(* Logix 5000 project; controller MV vendor 1 type 14 code 217 rev 31.11; software revision 31.00; part 30 of 53 *)
(* tags used below, declared in another part *)
   Alarm_Reset : BOOL;
   CWD : CHECKWORD_FLAGS;
   Default_Check_Time : DINT;
   Item_Faults_Are_Latched : BOOL;
   Item_Simulation_Flag : BOOL;
   MC_CH1_DR1 : PlantItem;   // CH1_DR1
   MC_CH1_DR1_ALARM : ALARM_DIGITAL;
   MC_CH1_DR1_C : ALIAS FOR RIO_Rack_2:4:I.Data.30;
   MC_CH1_DR1_DR : ALIAS FOR RIO_Rack_2:5:O.Data.14;
   MC_CH1_DR1_O : ALIAS FOR RIO_Rack_2:4:I.Data.26;
   MC_CH1_DR2 : PlantItem;   // CH1_DR2
   MC_CH1_DR2_ALARM : ALARM_DIGITAL;
   MC_CH1_DR2_C : ALIAS FOR RIO_Rack_2:4:I.Data.31;
   MC_CH1_DR2_DR : ALIAS FOR RIO_Rack_2:5:O.Data.15;
   MC_CH1_DR2_O : ALIAS FOR RIO_Rack_2:4:I.Data.27;
   MC_CH1_DRAIN : PlantItem;   // CH1_DRAIN
   MC_CH1_DRAIN_ALARM : ALARM_DIGITAL;
   MC_CH1_DRAIN_C : ALIAS FOR RIO_Rack_2:4:I.Data.28;
   MC_CH1_DRAIN_DR : ALIAS FOR RIO_Rack_2:5:O.Data.12;
   MC_CH1_DRAIN_O : ALIAS FOR RIO_Rack_2:4:I.Data.24;
   MC_CH1_DT1 : PlantItem;   // CH1_DT1
   MC_CH1_DT1_ALARM : ALARM_DIGITAL;
   MC_CH1_DT1_C : ALIAS FOR RIO_Rack_2:6:I.Data.4;
   MC_CH1_DT1_DR : ALIAS FOR RIO_Rack_2:5:O.Data.16;
   MC_CH1_DT1_O : ALIAS FOR RIO_Rack_2:6:I.Data.0;
   MC_CH1_DT2 : PlantItem;   // CH1_DT2
   MC_CH1_DT2_ALARM : ALARM_DIGITAL;
   MC_CH1_DT2_C : ALIAS FOR RIO_Rack_2:6:I.Data.5;
   MC_CH1_DT2_DR : ALIAS FOR RIO_Rack_2:5:O.Data.17;
   MC_CH1_DT2_O : ALIAS FOR RIO_Rack_2:6:I.Data.1;
   MC_CH1_LF1 : PlantItem;   // CH1_LF1
   MC_CH1_LF1_ALARM : ALARM_DIGITAL;
   MC_CH1_LF1_C : ALIAS FOR RIO_Rack_2:6:I.Data.7;
   MC_CH1_LF1_DR : ALIAS FOR RIO_Rack_2:5:O.Data.19;
   MC_CH1_LF1_O : ALIAS FOR RIO_Rack_2:6:I.Data.3;
   MC_CH1_PR1 : PlantItem;   // CH1_PR1
   MC_CH1_PR1_ALARM : ALARM_DIGITAL;
   MC_CH1_PR1_C : ALIAS FOR RIO_Rack_2:6:I.Data.6;
   MC_CH1_PR1_DR : ALIAS FOR RIO_Rack_2:5:O.Data.18;
   MC_CH1_PR1_O : ALIAS FOR RIO_Rack_2:6:I.Data.2;
   MC_CH1_R2R : PlantItem;   // CH1_R2R
   MC_CH1_R2R_ALARM : ALARM_DIGITAL;
   MC_CH1_R2R_C : ALIAS FOR RIO_Rack_2:4:I.Data.15;
   MC_CH1_R2R_DR : ALIAS FOR RIO_Rack_2:5:O.Data.7;
   MC_CH1_R2R_O : ALIAS FOR RIO_Rack_2:4:I.Data.11;
   MC_CH1_R3R : PlantItem;   // CH1_R3R
   MC_CH1_R3R_ALARM : ALARM_DIGITAL;
   MC_CH1_R3R_C : ALIAS FOR RIO_Rack_2:4:I.Data.20;
   MC_CH1_R3R_DR : ALIAS FOR RIO_Rack_2:5:O.Data.8;
   MC_CH1_R3R_O : ALIAS FOR RIO_Rack_2:4:I.Data.16;
   MC_CH1_R4R : PlantItem;   // CH1_R4R
   MC_CH1_R4R_ALARM : ALARM_DIGITAL;
   MC_CH1_R4R_C : ALIAS FOR RIO_Rack_2:4:I.Data.21;
   MC_CH1_R4R_DR : ALIAS FOR RIO_Rack_2:5:O.Data.9;
   MC_CH1_R4R_O : ALIAS FOR RIO_Rack_2:4:I.Data.17;
   MC_CH1_R5R : PlantItem;   // CH1_R5R
   MC_CH1_R5R_ALARM : ALARM_DIGITAL;
   MC_CH1_R5R_C : ALIAS FOR RIO_Rack_2:4:I.Data.22;
   MC_CH1_R5R_DR : ALIAS FOR RIO_Rack_2:5:O.Data.10;
   MC_CH1_R5R_O : ALIAS FOR RIO_Rack_2:4:I.Data.18;
   MC_CH1_R6R : PlantItem;   // CH1_R6R
   MC_CH1_R6R_ALARM : ALARM_DIGITAL;
   MC_CH1_R6R_C : ALIAS FOR RIO_Rack_2:4:I.Data.23;
   MC_CH1_R6R_DR : ALIAS FOR RIO_Rack_2:5:O.Data.11;
   MC_CH1_R6R_O : ALIAS FOR RIO_Rack_2:4:I.Data.19;
   MC_CH1_RR : PlantItem;   // CH1_RR
   MC_CH1_RR_ALARM : ALARM_DIGITAL;
   MC_CH1_RR_C : ALIAS FOR RIO_Rack_2:4:I.Data.29;
   MC_CH1_RR_DR : ALIAS FOR RIO_Rack_2:5:O.Data.13;
   MC_CH1_RR_O : ALIAS FOR RIO_Rack_2:4:I.Data.25;
   MC_CH2_R1 : PlantItem;   // CH2_R1
   MC_CH2_R1_ALARM : ALARM_DIGITAL;
   MC_CH2_R1_C : ALIAS FOR RIO_Rack_2:6:I.Data.12;
   MC_CH2_R1_DR : ALIAS FOR RIO_Rack_2:5:O.Data.20;
   MC_CH2_R1_O : ALIAS FOR RIO_Rack_2:6:I.Data.8;
   MC_CH2_R1R : PlantItem;   // CH2_R1R
   MC_CH2_R1R_ALARM : ALARM_DIGITAL;
   MC_CH2_R1R_C : ALIAS FOR RIO_Rack_2:6:I.Data.22;
   MC_CH2_R1R_DR : ALIAS FOR RIO_Rack_2:5:O.Data.26;
   MC_CH2_R1R_O : ALIAS FOR RIO_Rack_2:6:I.Data.18;
   MC_CH2_R2 : PlantItem;   // CH2_R2
   MC_CH2_R2_ALARM : ALARM_DIGITAL;
   MC_CH2_R2_C : ALIAS FOR RIO_Rack_2:6:I.Data.13;
   MC_CH2_R2_DR : ALIAS FOR RIO_Rack_2:5:O.Data.21;
   MC_CH2_R2_O : ALIAS FOR RIO_Rack_2:6:I.Data.9;
   MC_CH2_R2R : PlantItem;   // CH2_R2R
   MC_CH2_R2R_ALARM : ALARM_DIGITAL;
   MC_CH2_R2R_C : ALIAS FOR RIO_Rack_2:6:I.Data.23;
   MC_CH2_R2R_DR : ALIAS FOR RIO_Rack_2:5:O.Data.27;
   MC_CH2_R2R_O : ALIAS FOR RIO_Rack_2:6:I.Data.19;
   MC_CH2_R3 : PlantItem;   // CH2_R3
   MC_CH2_R3_ALARM : ALARM_DIGITAL;
   MC_CH2_R3_C : ALIAS FOR RIO_Rack_2:6:I.Data.14;
   MC_CH2_R3_DR : ALIAS FOR RIO_Rack_2:5:O.Data.22;
   MC_CH2_R3_O : ALIAS FOR RIO_Rack_2:6:I.Data.10;
   MC_CH2_R3R : PlantItem;   // CH2_R3R
   MC_CH2_R3R_ALARM : ALARM_DIGITAL;
   MC_CH2_R3R_C : ALIAS FOR RIO_Rack_2:6:I.Data.28;
   MC_CH2_R3R_DR : ALIAS FOR RIO_Rack_2:5:O.Data.28;
   MC_CH2_R3R_O : ALIAS FOR RIO_Rack_2:6:I.Data.24;
   MC_CH2_R4 : PlantItem;   // CH2_R4
   MC_CH2_R4_ALARM : ALARM_DIGITAL;
   MC_CH2_R4_C : ALIAS FOR RIO_Rack_2:6:I.Data.15;
   MC_CH2_R4_DR : ALIAS FOR RIO_Rack_2:5:O.Data.23;
   MC_CH2_R4_O : ALIAS FOR RIO_Rack_2:6:I.Data.11;
   MC_CH2_R4R : PlantItem;   // CH2_R4R
   MC_CH2_R4R_ALARM : ALARM_DIGITAL;
   MC_CH2_R4R_C : ALIAS FOR RIO_Rack_2:6:I.Data.29;
   MC_CH2_R4R_DR : ALIAS FOR RIO_Rack_2:5:O.Data.29;
   MC_CH2_R4R_O : ALIAS FOR RIO_Rack_2:6:I.Data.25;
   MC_CH2_R5 : PlantItem;   // CH2_R5
   MC_CH2_R5_ALARM : ALARM_DIGITAL;
   MC_CH2_R5_C : ALIAS FOR RIO_Rack_2:6:I.Data.20;
   MC_CH2_R5_DR : ALIAS FOR RIO_Rack_2:5:O.Data.24;
   MC_CH2_R5_O : ALIAS FOR RIO_Rack_2:6:I.Data.16;
   MC_CH2_R5R : PlantItem;   // CH2_R5R
   MC_CH2_R5R_ALARM : ALARM_DIGITAL;
   MC_CH2_R5R_C : ALIAS FOR RIO_Rack_2:6:I.Data.30;
   MC_CH2_R5R_DR : ALIAS FOR RIO_Rack_2:5:O.Data.30;
   MC_CH2_R5R_O : ALIAS FOR RIO_Rack_2:6:I.Data.26;
   MC_CH2_R6 : PlantItem;   // CH2_R6
   MC_CH2_R6_ALARM : ALARM_DIGITAL;
   MC_CH2_R6_C : ALIAS FOR RIO_Rack_2:6:I.Data.21;
   MC_CH2_R6_DR : ALIAS FOR RIO_Rack_2:5:O.Data.25;
   MC_CH2_R6_O : ALIAS FOR RIO_Rack_2:6:I.Data.17;
   One_Second_One_Scan : ALIAS FOR One_Second_1_scan;
(* MC_Common, continued *)

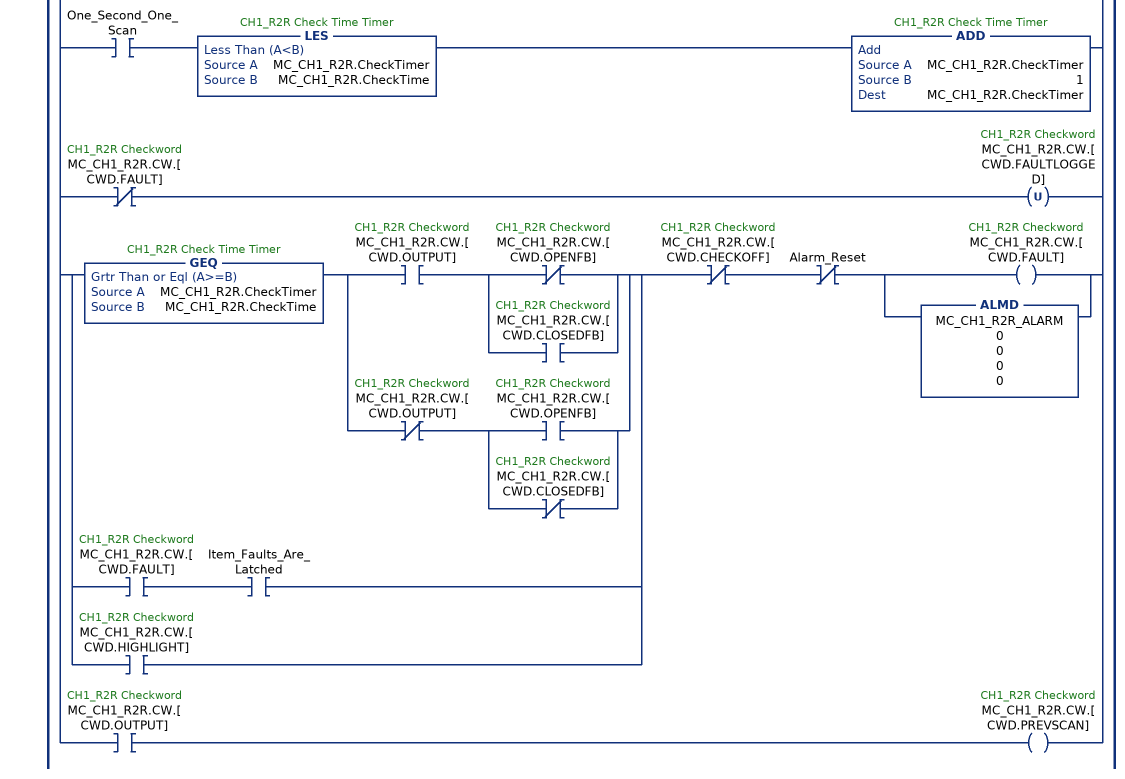
   [picture p611: MC_Common/MC_Valves rungs 7-7]
   7: [NEQ(MC_CH1_R2R.DriveBits,0) OTE(MC_CH1_R2R.CW.[CWD.AUTODRV]) ,[XIC(MC_CH1_R2R.CW.[CWD.AUTODRV]) XIO(MC_CH1_R2R.CW.[CWD.MANUAL]) ,XIC(MC_CH1_R2R.CW.[CWD.MANDRV]) XIC(MC_CH1_R2R.CW.[CWD.MANUAL]) ] OTE(MC_CH1_R2R.CW.[CWD.OUTPUT]) ,XIC(MC_CH1_R2R.CW.[CWD.OUTPUT]) OTE(MC_CH1_R2R_DR) ,XIC(S:FS) [OTU(MC_CH1_R2R.CW.[CWD.MANUAL]) ,LEQ(MC_CH1_R2R.CheckTime,0) MOV(Default_Check_Time,MC_CH1_R2R.CheckTime) ] ,[[XIC(MC_CH1_R2R_O) XIO(Item_Simulation_Flag) ,XIC(Item_Simulation_Flag) XIC(MC_CH1_R2R.CW.[CWD.OUTPUT]) XIO(MC_CH1_R2R.CW.[CWD.SIMFAIL]) ] OTE(MC_CH1_R2R.CW.[CWD.OPENFB]) ,[XIC(MC_CH1_R2R_C) XIO(Item_Simulation_Flag) ,XIC(Item_Simulation_Flag) XIO(MC_CH1_R2R.CW.[CWD.OUTPUT]) XIO(MC_CH1_R2R.CW.[CWD.SIMFAIL]) ] OTE(MC_CH1_R2R.CW.[CWD.CLOSEDFB]) ] ,[XIC(MC_CH1_R2R.CW.[CWD.OUTPUT]) XIO(MC_CH1_R2R.CW.[CWD.PREVSCAN]) ,XIO(MC_CH1_R2R.CW.[CWD.OUTPUT]) XIC(MC_CH1_R2R.CW.[CWD.PREVSCAN]) ] CLR(MC_CH1_R2R.CheckTimer) ,XIC(One_Second_One_Scan) LES(MC_CH1_R2R.CheckTimer,MC_CH1_R2R.CheckTime) ADD(MC_CH1_R2R.CheckTimer,1,MC_CH1_R2R.CheckTimer) ,XIO(MC_CH1_R2R.CW.[CWD.FAULT]) OTU(MC_CH1_R2R.CW.[CWD.FAULTLOGGED]) ,[GEQ(MC_CH1_R2R.CheckTimer,MC_CH1_R2R.CheckTime) [XIC(MC_CH1_R2R.CW.[CWD.OUTPUT]) [XIO(MC_CH1_R2R.CW.[CWD.OPENFB]) ,XIC(MC_CH1_R2R.CW.[CWD.CLOSEDFB]) ] ,XIO(MC_CH1_R2R.CW.[CWD.OUTPUT]) [XIC(MC_CH1_R2R.CW.[CWD.OPENFB]) ,XIO(MC_CH1_R2R.CW.[CWD.CLOSEDFB]) ] ] ,XIC(MC_CH1_R2R.CW.[CWD.FAULT]) XIC(Item_Faults_Are_Latched) ,XIC(MC_CH1_R2R.CW.[CWD.HIGHLIGHT]) ] XIO(MC_CH1_R2R.CW.[CWD.CHECKOFF]) XIO(Alarm_Reset) [OTE(MC_CH1_R2R.CW.[CWD.FAULT]) ,ALMD(MC_CH1_R2R_ALARM,0,0,0,0) ] ,XIC(MC_CH1_R2R.CW.[CWD.OUTPUT]) OTE(MC_CH1_R2R.CW.[CWD.PREVSCAN]) ];
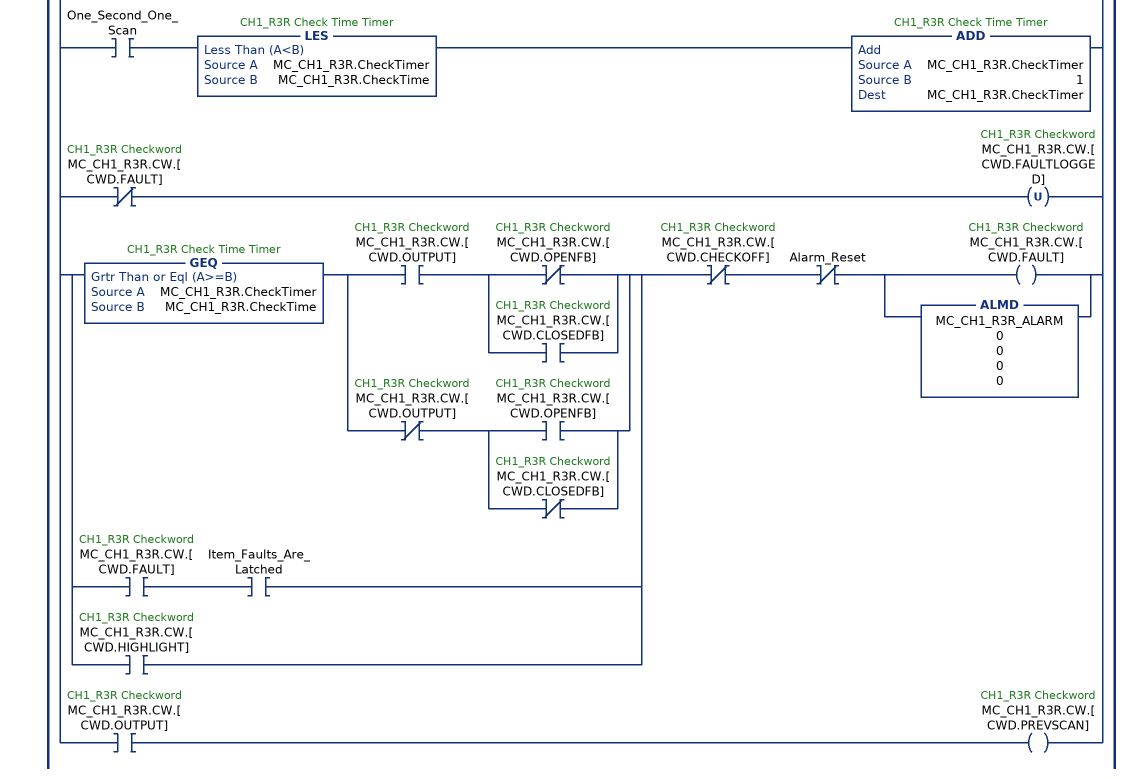
   8: [NEQ(MC_CH1_R3R.DriveBits,0) OTE(MC_CH1_R3R.CW.[CWD.AUTODRV]) ,[XIC(MC_CH1_R3R.CW.[CWD.AUTODRV]) XIO(MC_CH1_R3R.CW.[CWD.MANUAL]) ,XIC(MC_CH1_R3R.CW.[CWD.MANDRV]) XIC(MC_CH1_R3R.CW.[CWD.MANUAL]) ] OTE(MC_CH1_R3R.CW.[CWD.OUTPUT]) ,XIC(MC_CH1_R3R.CW.[CWD.OUTPUT]) OTE(MC_CH1_R3R_DR) ,XIC(S:FS) [OTU(MC_CH1_R3R.CW.[CWD.MANUAL]) ,LEQ(MC_CH1_R3R.CheckTime,0) MOV(Default_Check_Time,MC_CH1_R3R.CheckTime) ] ,[[XIC(MC_CH1_R3R_O) XIO(Item_Simulation_Flag) ,XIC(Item_Simulation_Flag) XIC(MC_CH1_R3R.CW.[CWD.OUTPUT]) XIO(MC_CH1_R3R.CW.[CWD.SIMFAIL]) ] OTE(MC_CH1_R3R.CW.[CWD.OPENFB]) ,[XIC(MC_CH1_R3R_C) XIO(Item_Simulation_Flag) ,XIC(Item_Simulation_Flag) XIO(MC_CH1_R3R.CW.[CWD.OUTPUT]) XIO(MC_CH1_R3R.CW.[CWD.SIMFAIL]) ] OTE(MC_CH1_R3R.CW.[CWD.CLOSEDFB]) ] ,[XIC(MC_CH1_R3R.CW.[CWD.OUTPUT]) XIO(MC_CH1_R3R.CW.[CWD.PREVSCAN]) ,XIO(MC_CH1_R3R.CW.[CWD.OUTPUT]) XIC(MC_CH1_R3R.CW.[CWD.PREVSCAN]) ] CLR(MC_CH1_R3R.CheckTimer) ,XIC(One_Second_One_Scan) LES(MC_CH1_R3R.CheckTimer,MC_CH1_R3R.CheckTime) ADD(MC_CH1_R3R.CheckTimer,1,MC_CH1_R3R.CheckTimer) ,XIO(MC_CH1_R3R.CW.[CWD.FAULT]) OTU(MC_CH1_R3R.CW.[CWD.FAULTLOGGED]) ,[GEQ(MC_CH1_R3R.CheckTimer,MC_CH1_R3R.CheckTime) [XIC(MC_CH1_R3R.CW.[CWD.OUTPUT]) [XIO(MC_CH1_R3R.CW.[CWD.OPENFB]) ,XIC(MC_CH1_R3R.CW.[CWD.CLOSEDFB]) ] ,XIO(MC_CH1_R3R.CW.[CWD.OUTPUT]) [XIC(MC_CH1_R3R.CW.[CWD.OPENFB]) ,XIO(MC_CH1_R3R.CW.[CWD.CLOSEDFB]) ] ] ,XIC(MC_CH1_R3R.CW.[CWD.FAULT]) XIC(Item_Faults_Are_Latched) ,XIC(MC_CH1_R3R.CW.[CWD.HIGHLIGHT]) ] XIO(MC_CH1_R3R.CW.[CWD.CHECKOFF]) XIO(Alarm_Reset) [OTE(MC_CH1_R3R.CW.[CWD.FAULT]) ,ALMD(MC_CH1_R3R_ALARM,0,0,0,0) ] ,XIC(MC_CH1_R3R.CW.[CWD.OUTPUT]) OTE(MC_CH1_R3R.CW.[CWD.PREVSCAN]) ];
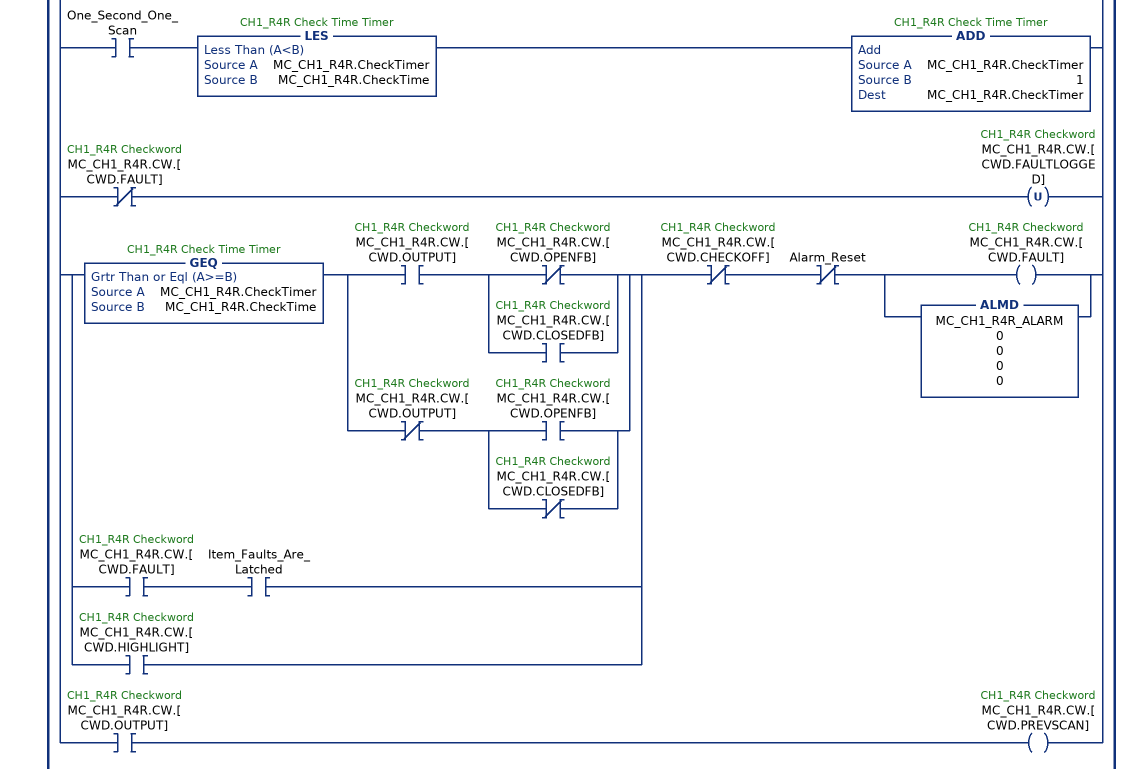
   9: [NEQ(MC_CH1_R4R.DriveBits,0) OTE(MC_CH1_R4R.CW.[CWD.AUTODRV]) ,[XIC(MC_CH1_R4R.CW.[CWD.AUTODRV]) XIO(MC_CH1_R4R.CW.[CWD.MANUAL]) ,XIC(MC_CH1_R4R.CW.[CWD.MANDRV]) XIC(MC_CH1_R4R.CW.[CWD.MANUAL]) ] OTE(MC_CH1_R4R.CW.[CWD.OUTPUT]) ,XIC(MC_CH1_R4R.CW.[CWD.OUTPUT]) OTE(MC_CH1_R4R_DR) ,XIC(S:FS) [OTU(MC_CH1_R4R.CW.[CWD.MANUAL]) ,LEQ(MC_CH1_R4R.CheckTime,0) MOV(Default_Check_Time,MC_CH1_R4R.CheckTime) ] ,[[XIC(MC_CH1_R4R_O) XIO(Item_Simulation_Flag) ,XIC(Item_Simulation_Flag) XIC(MC_CH1_R4R.CW.[CWD.OUTPUT]) XIO(MC_CH1_R4R.CW.[CWD.SIMFAIL]) ] OTE(MC_CH1_R4R.CW.[CWD.OPENFB]) ,[XIC(MC_CH1_R4R_C) XIO(Item_Simulation_Flag) ,XIC(Item_Simulation_Flag) XIO(MC_CH1_R4R.CW.[CWD.OUTPUT]) XIO(MC_CH1_R4R.CW.[CWD.SIMFAIL]) ] OTE(MC_CH1_R4R.CW.[CWD.CLOSEDFB]) ] ,[XIC(MC_CH1_R4R.CW.[CWD.OUTPUT]) XIO(MC_CH1_R4R.CW.[CWD.PREVSCAN]) ,XIO(MC_CH1_R4R.CW.[CWD.OUTPUT]) XIC(MC_CH1_R4R.CW.[CWD.PREVSCAN]) ] CLR(MC_CH1_R4R.CheckTimer) ,XIC(One_Second_One_Scan) LES(MC_CH1_R4R.CheckTimer,MC_CH1_R4R.CheckTime) ADD(MC_CH1_R4R.CheckTimer,1,MC_CH1_R4R.CheckTimer) ,XIO(MC_CH1_R4R.CW.[CWD.FAULT]) OTU(MC_CH1_R4R.CW.[CWD.FAULTLOGGED]) ,[GEQ(MC_CH1_R4R.CheckTimer,MC_CH1_R4R.CheckTime) [XIC(MC_CH1_R4R.CW.[CWD.OUTPUT]) [XIO(MC_CH1_R4R.CW.[CWD.OPENFB]) ,XIC(MC_CH1_R4R.CW.[CWD.CLOSEDFB]) ] ,XIO(MC_CH1_R4R.CW.[CWD.OUTPUT]) [XIC(MC_CH1_R4R.CW.[CWD.OPENFB]) ,XIO(MC_CH1_R4R.CW.[CWD.CLOSEDFB]) ] ] ,XIC(MC_CH1_R4R.CW.[CWD.FAULT]) XIC(Item_Faults_Are_Latched) ,XIC(MC_CH1_R4R.CW.[CWD.HIGHLIGHT]) ] XIO(MC_CH1_R4R.CW.[CWD.CHECKOFF]) XIO(Alarm_Reset) [OTE(MC_CH1_R4R.CW.[CWD.FAULT]) ,ALMD(MC_CH1_R4R_ALARM,0,0,0,0) ] ,XIC(MC_CH1_R4R.CW.[CWD.OUTPUT]) OTE(MC_CH1_R4R.CW.[CWD.PREVSCAN]) ];
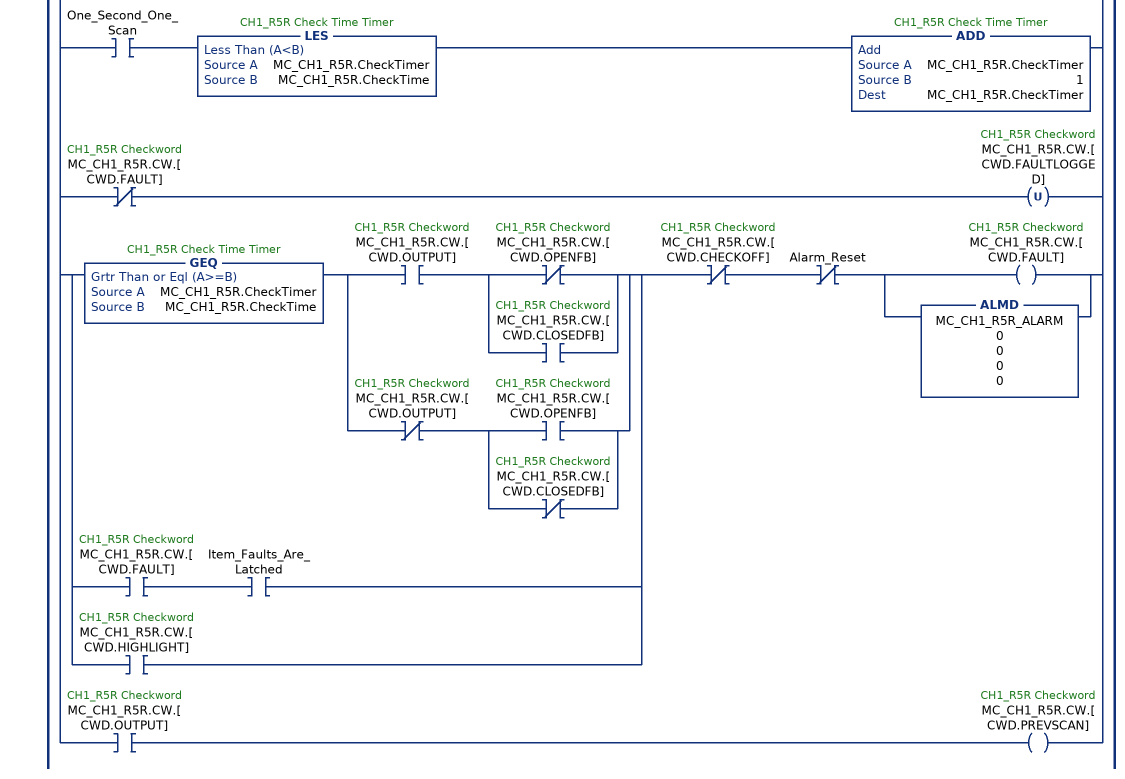
   10: [NEQ(MC_CH1_R5R.DriveBits,0) OTE(MC_CH1_R5R.CW.[CWD.AUTODRV]) ,[XIC(MC_CH1_R5R.CW.[CWD.AUTODRV]) XIO(MC_CH1_R5R.CW.[CWD.MANUAL]) ,XIC(MC_CH1_R5R.CW.[CWD.MANDRV]) XIC(MC_CH1_R5R.CW.[CWD.MANUAL]) ] OTE(MC_CH1_R5R.CW.[CWD.OUTPUT]) ,XIC(MC_CH1_R5R.CW.[CWD.OUTPUT]) OTE(MC_CH1_R5R_DR) ,XIC(S:FS) [OTU(MC_CH1_R5R.CW.[CWD.MANUAL]) ,LEQ(MC_CH1_R5R.CheckTime,0) MOV(Default_Check_Time,MC_CH1_R5R.CheckTime) ] ,[[XIC(MC_CH1_R5R_O) XIO(Item_Simulation_Flag) ,XIC(Item_Simulation_Flag) XIC(MC_CH1_R5R.CW.[CWD.OUTPUT]) XIO(MC_CH1_R5R.CW.[CWD.SIMFAIL]) ] OTE(MC_CH1_R5R.CW.[CWD.OPENFB]) ,[XIC(MC_CH1_R5R_C) XIO(Item_Simulation_Flag) ,XIC(Item_Simulation_Flag) XIO(MC_CH1_R5R.CW.[CWD.OUTPUT]) XIO(MC_CH1_R5R.CW.[CWD.SIMFAIL]) ] OTE(MC_CH1_R5R.CW.[CWD.CLOSEDFB]) ] ,[XIC(MC_CH1_R5R.CW.[CWD.OUTPUT]) XIO(MC_CH1_R5R.CW.[CWD.PREVSCAN]) ,XIO(MC_CH1_R5R.CW.[CWD.OUTPUT]) XIC(MC_CH1_R5R.CW.[CWD.PREVSCAN]) ] CLR(MC_CH1_R5R.CheckTimer) ,XIC(One_Second_One_Scan) LES(MC_CH1_R5R.CheckTimer,MC_CH1_R5R.CheckTime) ADD(MC_CH1_R5R.CheckTimer,1,MC_CH1_R5R.CheckTimer) ,XIO(MC_CH1_R5R.CW.[CWD.FAULT]) OTU(MC_CH1_R5R.CW.[CWD.FAULTLOGGED]) ,[GEQ(MC_CH1_R5R.CheckTimer,MC_CH1_R5R.CheckTime) [XIC(MC_CH1_R5R.CW.[CWD.OUTPUT]) [XIO(MC_CH1_R5R.CW.[CWD.OPENFB]) ,XIC(MC_CH1_R5R.CW.[CWD.CLOSEDFB]) ] ,XIO(MC_CH1_R5R.CW.[CWD.OUTPUT]) [XIC(MC_CH1_R5R.CW.[CWD.OPENFB]) ,XIO(MC_CH1_R5R.CW.[CWD.CLOSEDFB]) ] ] ,XIC(MC_CH1_R5R.CW.[CWD.FAULT]) XIC(Item_Faults_Are_Latched) ,XIC(MC_CH1_R5R.CW.[CWD.HIGHLIGHT]) ] XIO(MC_CH1_R5R.CW.[CWD.CHECKOFF]) XIO(Alarm_Reset) [OTE(MC_CH1_R5R.CW.[CWD.FAULT]) ,ALMD(MC_CH1_R5R_ALARM,0,0,0,0) ] ,XIC(MC_CH1_R5R.CW.[CWD.OUTPUT]) OTE(MC_CH1_R5R.CW.[CWD.PREVSCAN]) ];
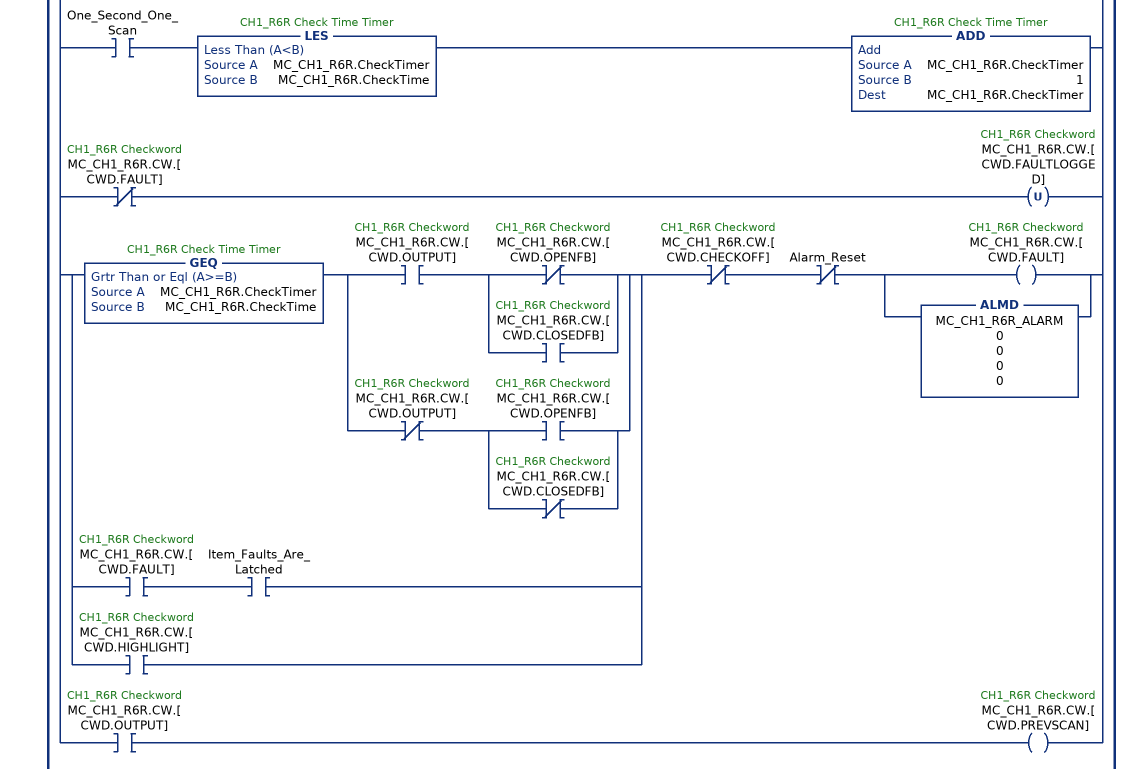
   11: [NEQ(MC_CH1_R6R.DriveBits,0) OTE(MC_CH1_R6R.CW.[CWD.AUTODRV]) ,[XIC(MC_CH1_R6R.CW.[CWD.AUTODRV]) XIO(MC_CH1_R6R.CW.[CWD.MANUAL]) ,XIC(MC_CH1_R6R.CW.[CWD.MANDRV]) XIC(MC_CH1_R6R.CW.[CWD.MANUAL]) ] OTE(MC_CH1_R6R.CW.[CWD.OUTPUT]) ,XIC(MC_CH1_R6R.CW.[CWD.OUTPUT]) OTE(MC_CH1_R6R_DR) ,XIC(S:FS) [OTU(MC_CH1_R6R.CW.[CWD.MANUAL]) ,LEQ(MC_CH1_R6R.CheckTime,0) MOV(Default_Check_Time,MC_CH1_R6R.CheckTime) ] ,[[XIC(MC_CH1_R6R_O) XIO(Item_Simulation_Flag) ,XIC(Item_Simulation_Flag) XIC(MC_CH1_R6R.CW.[CWD.OUTPUT]) XIO(MC_CH1_R6R.CW.[CWD.SIMFAIL]) ] OTE(MC_CH1_R6R.CW.[CWD.OPENFB]) ,[XIC(MC_CH1_R6R_C) XIO(Item_Simulation_Flag) ,XIC(Item_Simulation_Flag) XIO(MC_CH1_R6R.CW.[CWD.OUTPUT]) XIO(MC_CH1_R6R.CW.[CWD.SIMFAIL]) ] OTE(MC_CH1_R6R.CW.[CWD.CLOSEDFB]) ] ,[XIC(MC_CH1_R6R.CW.[CWD.OUTPUT]) XIO(MC_CH1_R6R.CW.[CWD.PREVSCAN]) ,XIO(MC_CH1_R6R.CW.[CWD.OUTPUT]) XIC(MC_CH1_R6R.CW.[CWD.PREVSCAN]) ] CLR(MC_CH1_R6R.CheckTimer) ,XIC(One_Second_One_Scan) LES(MC_CH1_R6R.CheckTimer,MC_CH1_R6R.CheckTime) ADD(MC_CH1_R6R.CheckTimer,1,MC_CH1_R6R.CheckTimer) ,XIO(MC_CH1_R6R.CW.[CWD.FAULT]) OTU(MC_CH1_R6R.CW.[CWD.FAULTLOGGED]) ,[GEQ(MC_CH1_R6R.CheckTimer,MC_CH1_R6R.CheckTime) [XIC(MC_CH1_R6R.CW.[CWD.OUTPUT]) [XIO(MC_CH1_R6R.CW.[CWD.OPENFB]) ,XIC(MC_CH1_R6R.CW.[CWD.CLOSEDFB]) ] ,XIO(MC_CH1_R6R.CW.[CWD.OUTPUT]) [XIC(MC_CH1_R6R.CW.[CWD.OPENFB]) ,XIO(MC_CH1_R6R.CW.[CWD.CLOSEDFB]) ] ] ,XIC(MC_CH1_R6R.CW.[CWD.FAULT]) XIC(Item_Faults_Are_Latched) ,XIC(MC_CH1_R6R.CW.[CWD.HIGHLIGHT]) ] XIO(MC_CH1_R6R.CW.[CWD.CHECKOFF]) XIO(Alarm_Reset) [OTE(MC_CH1_R6R.CW.[CWD.FAULT]) ,ALMD(MC_CH1_R6R_ALARM,0,0,0,0) ] ,XIC(MC_CH1_R6R.CW.[CWD.OUTPUT]) OTE(MC_CH1_R6R.CW.[CWD.PREVSCAN]) ];
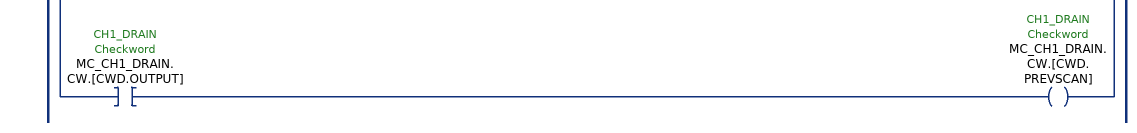
   12: [NEQ(MC_CH1_DRAIN.DriveBits,0) OTE(MC_CH1_DRAIN.CW.[CWD.AUTODRV]) ,[XIC(MC_CH1_DRAIN.CW.[CWD.AUTODRV]) XIO(MC_CH1_DRAIN.CW.[CWD.MANUAL]) ,XIC(MC_CH1_DRAIN.CW.[CWD.MANDRV]) XIC(MC_CH1_DRAIN.CW.[CWD.MANUAL]) ] OTE(MC_CH1_DRAIN.CW.[CWD.OUTPUT]) ,XIC(MC_CH1_DRAIN.CW.[CWD.OUTPUT]) OTE(MC_CH1_DRAIN_DR) ,XIC(S:FS) [OTU(MC_CH1_DRAIN.CW.[CWD.MANUAL]) ,LEQ(MC_CH1_DRAIN.CheckTime,0) MOV(Default_Check_Time,MC_CH1_DRAIN.CheckTime) ] ,[[XIC(MC_CH1_DRAIN_O) XIO(Item_Simulation_Flag) ,XIC(Item_Simulation_Flag) XIC(MC_CH1_DRAIN.CW.[CWD.OUTPUT]) XIO(MC_CH1_DRAIN.CW.[CWD.SIMFAIL]) ] OTE(MC_CH1_DRAIN.CW.[CWD.OPENFB]) ,[XIC(MC_CH1_DRAIN_C) XIO(Item_Simulation_Flag) ,XIC(Item_Simulation_Flag) XIO(MC_CH1_DRAIN.CW.[CWD.OUTPUT]) XIO(MC_CH1_DRAIN.CW.[CWD.SIMFAIL]) ] OTE(MC_CH1_DRAIN.CW.[CWD.CLOSEDFB]) ] ,[XIC(MC_CH1_DRAIN.CW.[CWD.OUTPUT]) XIO(MC_CH1_DRAIN.CW.[CWD.PREVSCAN]) ,XIO(MC_CH1_DRAIN.CW.[CWD.OUTPUT]) XIC(MC_CH1_DRAIN.CW.[CWD.PREVSCAN]) ] CLR(MC_CH1_DRAIN.CheckTimer) ,XIC(One_Second_One_Scan) LES(MC_CH1_DRAIN.CheckTimer,MC_CH1_DRAIN.CheckTime) ADD(MC_CH1_DRAIN.CheckTimer,1,MC_CH1_DRAIN.CheckTimer) ,XIO(MC_CH1_DRAIN.CW.[CWD.FAULT]) OTU(MC_CH1_DRAIN.CW.[CWD.FAULTLOGGED]) ,[GEQ(MC_CH1_DRAIN.CheckTimer,MC_CH1_DRAIN.CheckTime) [XIC(MC_CH1_DRAIN.CW.[CWD.OUTPUT]) [XIO(MC_CH1_DRAIN.CW.[CWD.OPENFB]) ,XIC(MC_CH1_DRAIN.CW.[CWD.CLOSEDFB]) ] ,XIO(MC_CH1_DRAIN.CW.[CWD.OUTPUT]) [XIC(MC_CH1_DRAIN.CW.[CWD.OPENFB]) ,XIO(MC_CH1_DRAIN.CW.[CWD.CLOSEDFB]) ] ] ,XIC(MC_CH1_DRAIN.CW.[CWD.FAULT]) XIC(Item_Faults_Are_Latched) ,XIC(MC_CH1_DRAIN.CW.[CWD.HIGHLIGHT]) ] XIO(MC_CH1_DRAIN.CW.[CWD.CHECKOFF]) XIO(Alarm_Reset) [OTE(MC_CH1_DRAIN.CW.[CWD.FAULT]) ,ALMD(MC_CH1_DRAIN_ALARM,0,0,0,0) ] ,XIC(MC_CH1_DRAIN.CW.[CWD.OUTPUT]) OTE(MC_CH1_DRAIN.CW.[CWD.PREVSCAN]) ];
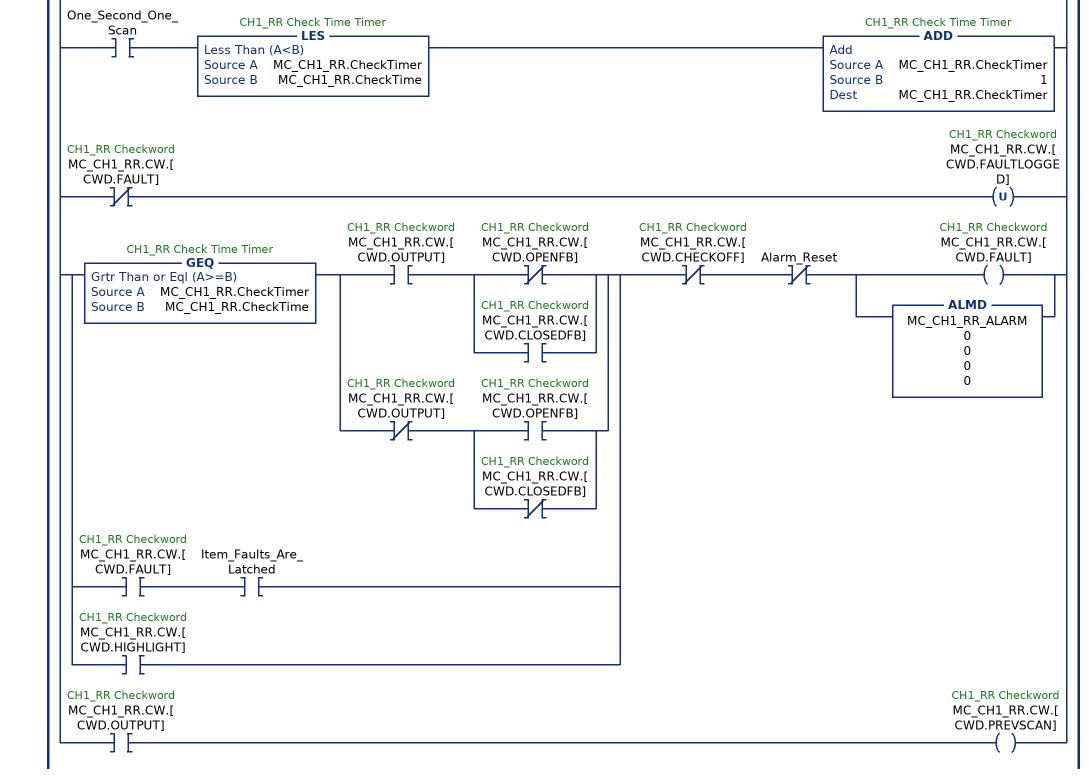
   13: [NEQ(MC_CH1_RR.DriveBits,0) OTE(MC_CH1_RR.CW.[CWD.AUTODRV]) ,[XIC(MC_CH1_RR.CW.[CWD.AUTODRV]) XIO(MC_CH1_RR.CW.[CWD.MANUAL]) ,XIC(MC_CH1_RR.CW.[CWD.MANDRV]) XIC(MC_CH1_RR.CW.[CWD.MANUAL]) ] OTE(MC_CH1_RR.CW.[CWD.OUTPUT]) ,XIC(MC_CH1_RR.CW.[CWD.OUTPUT]) OTE(MC_CH1_RR_DR) ,XIC(S:FS) [OTU(MC_CH1_RR.CW.[CWD.MANUAL]) ,LEQ(MC_CH1_RR.CheckTime,0) MOV(Default_Check_Time,MC_CH1_RR.CheckTime) ] ,[[XIC(MC_CH1_RR_O) XIO(Item_Simulation_Flag) ,XIC(Item_Simulation_Flag) XIC(MC_CH1_RR.CW.[CWD.OUTPUT]) XIO(MC_CH1_RR.CW.[CWD.SIMFAIL]) ] OTE(MC_CH1_RR.CW.[CWD.OPENFB]) ,[XIC(MC_CH1_RR_C) XIO(Item_Simulation_Flag) ,XIC(Item_Simulation_Flag) XIO(MC_CH1_RR.CW.[CWD.OUTPUT]) XIO(MC_CH1_RR.CW.[CWD.SIMFAIL]) ] OTE(MC_CH1_RR.CW.[CWD.CLOSEDFB]) ] ,[XIC(MC_CH1_RR.CW.[CWD.OUTPUT]) XIO(MC_CH1_RR.CW.[CWD.PREVSCAN]) ,XIO(MC_CH1_RR.CW.[CWD.OUTPUT]) XIC(MC_CH1_RR.CW.[CWD.PREVSCAN]) ] CLR(MC_CH1_RR.CheckTimer) ,XIC(One_Second_One_Scan) LES(MC_CH1_RR.CheckTimer,MC_CH1_RR.CheckTime) ADD(MC_CH1_RR.CheckTimer,1,MC_CH1_RR.CheckTimer) ,XIO(MC_CH1_RR.CW.[CWD.FAULT]) OTU(MC_CH1_RR.CW.[CWD.FAULTLOGGED]) ,[GEQ(MC_CH1_RR.CheckTimer,MC_CH1_RR.CheckTime) [XIC(MC_CH1_RR.CW.[CWD.OUTPUT]) [XIO(MC_CH1_RR.CW.[CWD.OPENFB]) ,XIC(MC_CH1_RR.CW.[CWD.CLOSEDFB]) ] ,XIO(MC_CH1_RR.CW.[CWD.OUTPUT]) [XIC(MC_CH1_RR.CW.[CWD.OPENFB]) ,XIO(MC_CH1_RR.CW.[CWD.CLOSEDFB]) ] ] ,XIC(MC_CH1_RR.CW.[CWD.FAULT]) XIC(Item_Faults_Are_Latched) ,XIC(MC_CH1_RR.CW.[CWD.HIGHLIGHT]) ] XIO(MC_CH1_RR.CW.[CWD.CHECKOFF]) XIO(Alarm_Reset) [OTE(MC_CH1_RR.CW.[CWD.FAULT]) ,ALMD(MC_CH1_RR_ALARM,0,0,0,0) ] ,XIC(MC_CH1_RR.CW.[CWD.OUTPUT]) OTE(MC_CH1_RR.CW.[CWD.PREVSCAN]) ];